// TIA Portal project "Network_1.0" (V15.1) (continued)
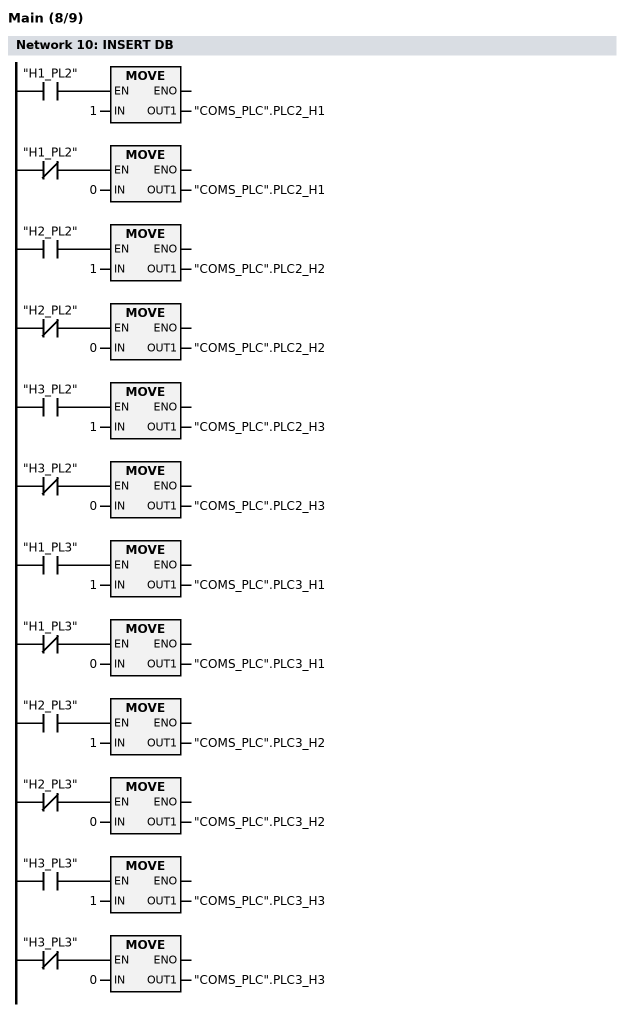
   RUNG wire#powerrail
      Contact( "H1_PL2" )
      Move(in := 1, out1 => "COMS_PLC".PLC2_H1)
   END_RUNG
   RUNG wire#powerrail
      I_Contact( "H1_PL2" )
      Move(in := 0, out1 => "COMS_PLC".PLC2_H1)
   END_RUNG
   RUNG wire#powerrail
      Contact( "H2_PL2" )
      Move(in := 1, out1 => "COMS_PLC".PLC2_H2)
   END_RUNG
   RUNG wire#powerrail
      I_Contact( "H2_PL2" )
      Move(in := 0, out1 => "COMS_PLC".PLC2_H2)
   END_RUNG
   RUNG wire#powerrail
      Contact( "H3_PL2" )
      Move(in := 1, out1 => "COMS_PLC".PLC2_H3)
   END_RUNG
   RUNG wire#powerrail
      I_Contact( "H3_PL2" )
      Move(in := 0, out1 => "COMS_PLC".PLC2_H3)
   END_RUNG
   RUNG wire#powerrail
      Contact( "H1_PL3" )
      Move(in := 1, out1 => "COMS_PLC".PLC3_H1)
   END_RUNG
   RUNG wire#powerrail
      I_Contact( "H1_PL3" )
      Move(in := 0, out1 => "COMS_PLC".PLC3_H1)
   END_RUNG
   RUNG wire#powerrail
      Contact( "H2_PL3" )
      Move(in := 1, out1 => "COMS_PLC".PLC3_H2)
   END_RUNG
   RUNG wire#powerrail
      I_Contact( "H2_PL3" )
      Move(in := 0, out1 => "COMS_PLC".PLC3_H2)
   END_RUNG
   RUNG wire#powerrail
      Contact( "H3_PL3" )
      Move(in := 1, out1 => "COMS_PLC".PLC3_H3)
   END_RUNG
   RUNG wire#powerrail
      I_Contact( "H3_PL3" )
      Move(in := 0, out1 => "COMS_PLC".PLC3_H3)
   END_RUNG
   // the same network as SCL:
   IF "H1_PL2" THEN "COMS_PLC".PLC2_H1 := 1; END_IF;
   IF NOT "H1_PL2" THEN "COMS_PLC".PLC2_H1 := 0; END_IF;
   IF "H2_PL2" THEN "COMS_PLC".PLC2_H2 := 1; END_IF;
   IF NOT "H2_PL2" THEN "COMS_PLC".PLC2_H2 := 0; END_IF;
   IF "H3_PL2" THEN "COMS_PLC".PLC2_H3 := 1; END_IF;
   IF NOT "H3_PL2" THEN "COMS_PLC".PLC2_H3 := 0; END_IF;
   IF "H1_PL3" THEN "COMS_PLC".PLC3_H1 := 1; END_IF;
   IF NOT "H1_PL3" THEN "COMS_PLC".PLC3_H1 := 0; END_IF;
   IF "H2_PL3" THEN "COMS_PLC".PLC3_H2 := 1; END_IF;
   IF NOT "H2_PL3" THEN "COMS_PLC".PLC3_H2 := 0; END_IF;
   IF "H3_PL3" THEN "COMS_PLC".PLC3_H3 := 1; END_IF;
   IF NOT "H3_PL3" THEN "COMS_PLC".PLC3_H3 := 0; END_IF;
END_REGION

REGION Network 11: GET
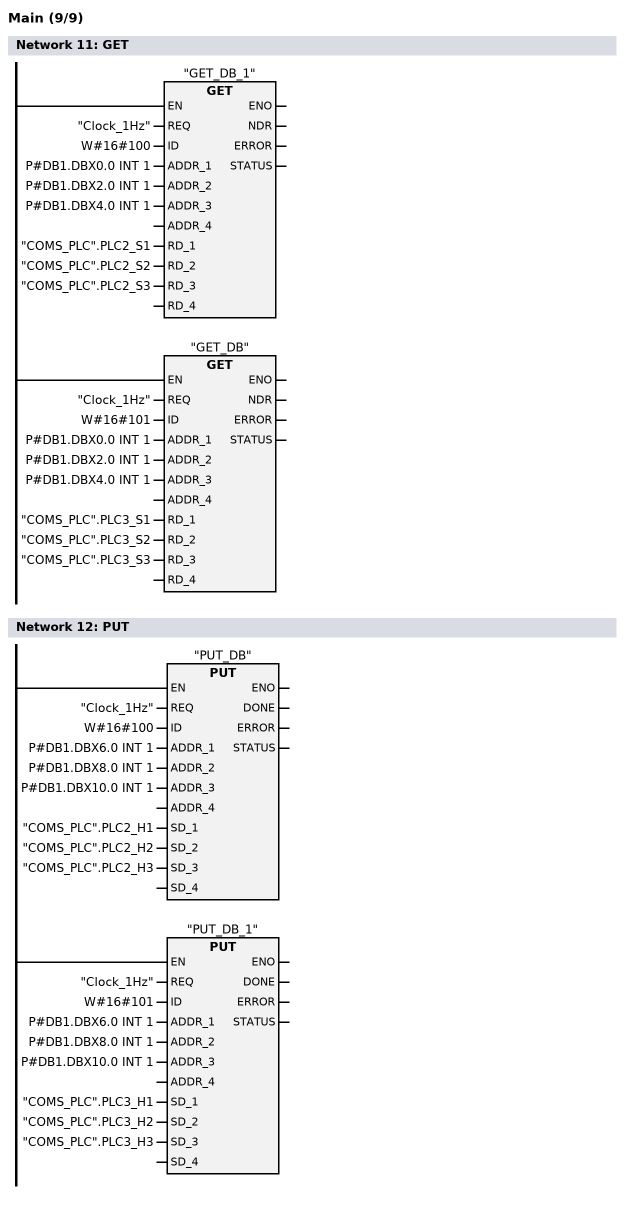
   "GET_DB_1"(REQ := "Clock_1Hz",   // GET
              ID := W#16#100,
              ADDR_1 := P#DB1.DBX0.0 INT 1,
              ADDR_2 := P#DB1.DBX2.0 INT 1,
              ADDR_3 := P#DB1.DBX4.0 INT 1,
              RD_1 := "COMS_PLC".PLC2_S1,
              RD_2 := "COMS_PLC".PLC2_S2,
              RD_3 := "COMS_PLC".PLC2_S3);
   "GET_DB"(REQ := "Clock_1Hz",   // GET
            ID := W#16#101,
            ADDR_1 := P#DB1.DBX0.0 INT 1,
            ADDR_2 := P#DB1.DBX2.0 INT 1,
            ADDR_3 := P#DB1.DBX4.0 INT 1,
            RD_1 := "COMS_PLC".PLC3_S1,
            RD_2 := "COMS_PLC".PLC3_S2,
            RD_3 := "COMS_PLC".PLC3_S3);
END_REGION

REGION Network 12: PUT
   "PUT_DB"(REQ := "Clock_1Hz",   // PUT
            ID := W#16#100,
            ADDR_1 := P#DB1.DBX6.0 INT 1,
            ADDR_2 := P#DB1.DBX8.0 INT 1,
            ADDR_3 := P#DB1.DBX10.0 INT 1,
            SD_1 := "COMS_PLC".PLC2_H1,
            SD_2 := "COMS_PLC".PLC2_H2,
            SD_3 := "COMS_PLC".PLC2_H3);
   "PUT_DB_1"(REQ := "Clock_1Hz",   // PUT
              ID := W#16#101,
              ADDR_1 := P#DB1.DBX6.0 INT 1,
              ADDR_2 := P#DB1.DBX8.0 INT 1,
              ADDR_3 := P#DB1.DBX10.0 INT 1,
              SD_1 := "COMS_PLC".PLC3_H1,
              SD_2 := "COMS_PLC".PLC3_H2,
              SD_3 := "COMS_PLC".PLC3_H3);
END_REGION
END_ORGANIZATION_BLOCK

// ===== PLC "PLC_2"  CPU 1215C DC/DC/DC =====

VAR_GLOBAL   // PLC tag table "Default tag table"
   "S4_JR" AT %I0.0 : Bool;
   "S3_JR" AT %I0.1 : Bool;
   "H2_JR" AT %Q0.1 : Bool;
   "S2_JR" AT %I0.2 : Bool;
   "S1_JR" AT %I0.3 : Bool;
   "PE_JR" AT %I0.4 : Bool;
   "H1_JR" AT %Q0.2 : Bool;
   "H3_JR" AT %Q0.0 : Bool;
   "Clock_Byte" AT %MB0 : Byte;
   "Clock_10Hz" AT %M0.0 : Bool;
   "Clock_5Hz" AT %M0.1 : Bool;
   "Clock_2.5Hz" AT %M0.2 : Bool;
   "Clock_2Hz" AT %M0.3 : Bool;
   "Clock_1.25Hz" AT %M0.4 : Bool;
   "Clock_1Hz" AT %M0.5 : Bool;
   "Clock_0.625Hz" AT %M0.6 : Bool;
   "Clock_0.5Hz" AT %M0.7 : Bool;
END_VAR

VAR_GLOBAL CONSTANT   // PLC tag table "Default tag table"
   "PLC_2" : Byte := 11;   // 2
END_VAR

DATA_BLOCK "Prueba"   // DB1
{ S7_Optimized_Access := 'FALSE' }
VERSION : 0.1
   VAR
      S1 : Int;
      S2 : Int;
      S3 : Int;
      H1 : Int;
      H2 : Int;
      H3 : Int;
   END_VAR
BEGIN
END_DATA_BLOCK

ORGANIZATION_BLOCK "Main"   // OB1, LAD, ProgramCycle
TITLE = "Main Program Sweep (Cycle)"
{ S7_Optimized_Access := 'TRUE' }
VERSION : 0.1
   VAR_INPUT
      Initial_Call : Bool;   // Initial call of this OB
      Remanence : Bool;   // =True, if remanent data are available
   END_VAR
BEGIN

REGION Network 1: SET DB
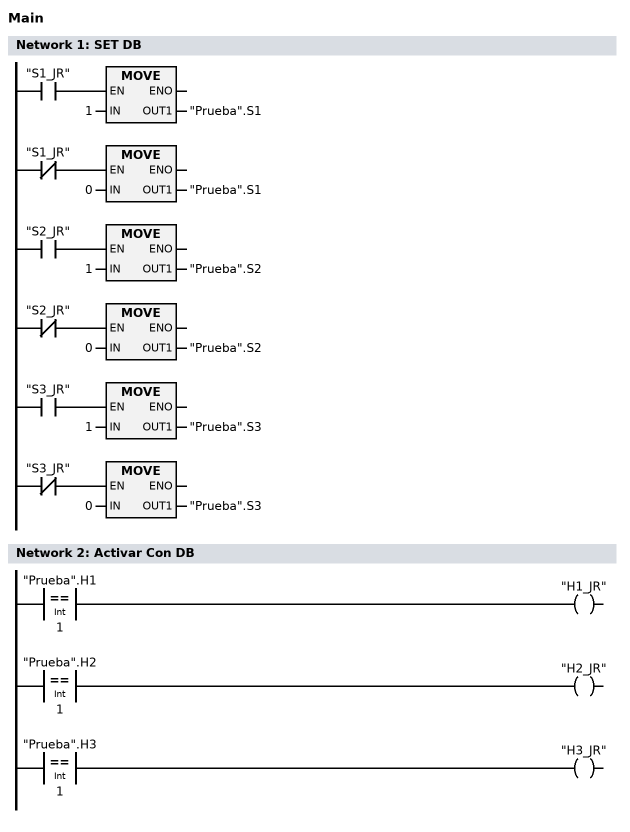
   RUNG wire#powerrail
      Contact( "S1_JR" )
      Move(in := 1, out1 => "Prueba".S1)
   END_RUNG
   RUNG wire#powerrail
      I_Contact( "S1_JR" )
      Move(in := 0, out1 => "Prueba".S1)
   END_RUNG
   RUNG wire#powerrail
      Contact( "S2_JR" )
      Move(in := 1, out1 => "Prueba".S2)
   END_RUNG
   RUNG wire#powerrail
      I_Contact( "S2_JR" )
      Move(in := 0, out1 => "Prueba".S2)
   END_RUNG
   RUNG wire#powerrail
      Contact( "S3_JR" )
      Move(in := 1, out1 => "Prueba".S3)
   END_RUNG
   RUNG wire#powerrail
      I_Contact( "S3_JR" )
      Move(in := 0, out1 => "Prueba".S3)
   END_RUNG
   // the same network as SCL:
   IF "S1_JR" THEN "Prueba".S1 := 1; END_IF;
   IF NOT "S1_JR" THEN "Prueba".S1 := 0; END_IF;
   IF "S2_JR" THEN "Prueba".S2 := 1; END_IF;
   IF NOT "S2_JR" THEN "Prueba".S2 := 0; END_IF;
   IF "S3_JR" THEN "Prueba".S3 := 1; END_IF;
   IF NOT "S3_JR" THEN "Prueba".S3 := 0; END_IF;
END_REGION

REGION Network 2: Activar Con DB
   RUNG wire#powerrail
      { S7_Templates := "SrcType := Int" } EQ_Contact(in1 := "Prueba".H1, in2 := 1)
      Coil( "H1_JR" )
   END_RUNG
   RUNG wire#powerrail
      { S7_Templates := "SrcType := Int" } EQ_Contact(in1 := "Prueba".H2, in2 := 1)
      Coil( "H2_JR" )
   END_RUNG
   RUNG wire#powerrail
      { S7_Templates := "SrcType := Int" } EQ_Contact(in1 := "Prueba".H3, in2 := 1)
      Coil( "H3_JR" )
   END_RUNG
   // the same network as SCL:
   "H1_JR" := "Prueba".H1 = 1;
   "H2_JR" := "Prueba".H2 = 1;
   "H3_JR" := "Prueba".H3 = 1;
END_REGION
END_ORGANIZATION_BLOCK

// ===== PLC "PLC_3"  CPU 1215C DC/DC/DC =====

VAR_GLOBAL   // PLC tag table "Default tag table"
   "H1_FE" AT %Q0.0 : Bool;
   "PE_FE" AT %I0.0 : Bool;
   "S1_FE" AT %I0.1 : Bool;
   "S2_FE" AT %I0.2 : Bool;
   "S3_FE" AT %I0.3 : Bool;
   "H2_FE" AT %Q0.1 : Bool;
   "H3_FE" AT %Q0.2 : Bool;
END_VAR

DATA_BLOCK "Control_PLC3"   // DB1
{ S7_Optimized_Access := 'FALSE' }
VERSION : 0.1
   VAR
      S1 : Int;
      S2 : Int;
      S3 : Int;
      H1 : Int;
      H2 : Int;
      H3 : Int;
   END_VAR
BEGIN
END_DATA_BLOCK

ORGANIZATION_BLOCK "Main"   // OB1, LAD, ProgramCycle
TITLE = "Main Program Sweep (Cycle)"
{ S7_Optimized_Access := 'TRUE' }
VERSION : 0.1
   VAR_INPUT
      Initial_Call : Bool;   // Initial call of this OB
      Remanence : Bool;   // =True, if remanent data are available
   END_VAR
BEGIN

REGION Network 1: SET DB
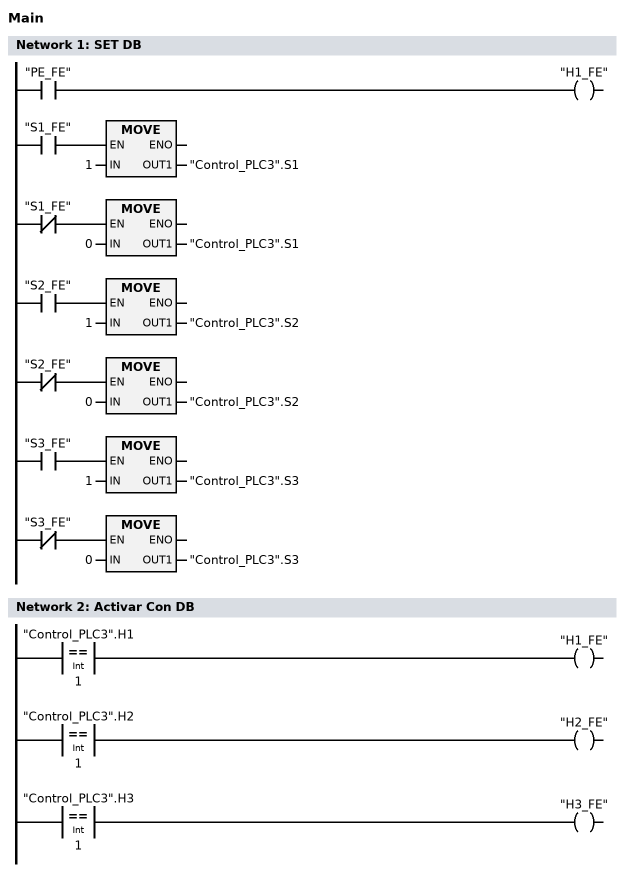
   RUNG wire#powerrail
      Contact( "PE_FE" )
      Coil( "H1_FE" )
   END_RUNG
   RUNG wire#powerrail
      Contact( "S1_FE" )
      Move(in := 1, out1 => "Control_PLC3".S1)
   END_RUNG
   RUNG wire#powerrail
      I_Contact( "S1_FE" )
      Move(in := 0, out1 => "Control_PLC3".S1)
   END_RUNG
   RUNG wire#powerrail
      Contact( "S2_FE" )
      Move(in := 1, out1 => "Control_PLC3".S2)
   END_RUNG
   RUNG wire#powerrail
      I_Contact( "S2_FE" )
      Move(in := 0, out1 => "Control_PLC3".S2)
   END_RUNG
   RUNG wire#powerrail
      Contact( "S3_FE" )
      Move(in := 1, out1 => "Control_PLC3".S3)
   END_RUNG
   RUNG wire#powerrail
      I_Contact( "S3_FE" )
      Move(in := 0, out1 => "Control_PLC3".S3)
   END_RUNG
   // the same network as SCL:
   "H1_FE" := "PE_FE";
   IF "S1_FE" THEN "Control_PLC3".S1 := 1; END_IF;
   IF NOT "S1_FE" THEN "Control_PLC3".S1 := 0; END_IF;
   IF "S2_FE" THEN "Control_PLC3".S2 := 1; END_IF;
   IF NOT "S2_FE" THEN "Control_PLC3".S2 := 0; END_IF;
   IF "S3_FE" THEN "Control_PLC3".S3 := 1; END_IF;
   IF NOT "S3_FE" THEN "Control_PLC3".S3 := 0; END_IF;
END_REGION

REGION Network 2: Activar Con DB
   RUNG wire#powerrail
      { S7_Templates := "SrcType := Int" } EQ_Contact(in1 := "Control_PLC3".H1, in2 := 1)
      Coil( "H1_FE" )
   END_RUNG
   RUNG wire#powerrail
      { S7_Templates := "SrcType := Int" } EQ_Contact(in1 := "Control_PLC3".H2, in2 := 1)
      Coil( "H2_FE" )
   END_RUNG
   RUNG wire#powerrail
      { S7_Templates := "SrcType := Int" } EQ_Contact(in1 := "Control_PLC3".H3, in2 := 1)
      Coil( "H3_FE" )
   END_RUNG
   // the same network as SCL:
   "H1_FE" := "Control_PLC3".H1 = 1;
   "H2_FE" := "Control_PLC3".H2 = 1;
   "H3_FE" := "Control_PLC3".H3 = 1;
END_REGION
END_ORGANIZATION_BLOCK

(* ===== HMI "HMI_RT_1" =====
system functions are stored by id; their names below are inferred from use
connection "HMI_Connection_1": ETHERNET, SMART_S7_1500_OMS

HMI tags "Default tag table"
   "Tag_ScreenNumber" : UInt, internal
   "S1" : Bool = PLC S1_HM1 AT %M3.0, 100 ms
   "S2" : Bool = PLC S2_HM1 AT %M3.1, 100 ms
   "S3" : Bool = PLC S3_HM1 AT %M3.2, 100 ms
   "H1_HM1" : Bool = PLC H1_HM1 AT %M6.3, 100 ms
   "H2_HM1" : Bool = PLC H2_HM1 AT %M6.4, 100 ms
   "H3_HM1" : Bool = PLC H3_HM1 AT %M6.5, 100 ms
   "Selector" : UInt = PLC Selector_HMI_1 AT %MW8, 100 ms

text list "PLC_SELECTOR": 1 'Betsy'; 2 'JR'; 3 'Fer'

Template "Template_1" 480x272
   Button "Exit" at 388,227 size 63x44; TextOff 'Exit'; PictureOff "ExitRuntime_KTP400_Basic_PN_TR"; PictureOn "ExitRuntime_KTP400_Basic_PN_TR"
      on Release: StopRuntime(0)
   Button "Log on" at 268,227 size 63x44; TextOff 'Log on'; PictureOff "Login_KTP400_Basic_PN_TR"; PictureOn "Login_KTP400_Basic_PN_TR"
      on Release: function_a2a04561()
   Button "Alarms" at 148,227 size 63x44; TextOff 'Alarms'; PictureOff "AlarmDisplay_KTP400_Basic_PN_TR"; PictureOn "AlarmDisplay_KTP400_Basic_PN_TR"
      on Release: function_ef3f5d25("Alarm window_Unacknowledged", -1)
   Button "Start screen" at 28,227 size 63x44; TextOff 'Start screen'; PictureOff "NavigateHome_KTP400_Basic_PN_TR"; PictureOn "NavigateHome_KTP400_Basic_PN_TR"
      on Release: ActivateScreen("Root screen", 0)
   SymbolicIOField "Symbolic_IO_Field_Screen" at 162,8 size 231x29; TextOff '0'; TextOn '1'; TextList "TextList_ScreenNames"
      ProcessValue <- "Tag_ScreenNumber"
      on Change: ActivateScreenByNumber("Tag_ScreenNumber", 0)
   DateTimeField "HmiScreenItemData" at 395,22 size 85x22
   DateTimeField "HmiScreenItemData_1" at 395,0 size 85x22
   GraphicView "Logo" at 0,0 size 160x45; Picture "Logo of HMI_1"

screen "Root screen" 480x272, template "Template_1"
   on GenerateScreen: SetTag("Tag_ScreenNumber", 1)
   Button "Button_1" at 169,112 size 146x61; TextOff 'LED CONTROL'
      on Click: ActivateScreen("Led_control", 8)

screen "SIMATIC PLC system diagnostics" 480x272, template "Template_1"
   on GenerateScreen: SetTag("Tag_ScreenNumber", 3)
   SysDiagControl "HmiScreenItemData" at 1,77 size 476x143
   Button "Back" at 1,46 size 157x30; TextOff 'Back'
      on Release: ActivateScreen("Root screen", 0)

screen "Project information" 480x272, template "Template_1"
   on GenerateScreen: SetTag("Tag_ScreenNumber", 4)
   TextField "HmiScreenItemData" at 4,78 size 184x20; Text 'Project name:'
   TextField "HmiScreenItemData_1" at 192,78 size 284x20; Text 'Network_1'
   TextField "HmiScreenItemData_2" at 4,99 size 184x20; Text 'Created on:'
   TextField "HmiScreenItemData_3" at 192,99 size 284x20; Text '3/10/2025 2:35:17 PM'
   TextField "HmiScreenItemData_4" at 4,120 size 184x20; Text 'Author:'
   TextField "HmiScreenItemData_5" at 192,120 size 284x20; Text '192072'
   TextField "HmiScreenItemData_6" at 4,141 size 184x20; Text 'Description:'
   TextField "HmiScreenItemData_7" at 192,141 size 284x20; Text '(not configured)'
   Button "Back" at 1,46 size 157x30; TextOff 'Back'
      on Release: ActivateScreen("Root screen", 0)

screen "System information" 480x272, template "Template_1"
   on GenerateScreen: SetTag("Tag_ScreenNumber", 6)
   TextField "HmiScreenItemData" at 4,78 size 184x20; Text 'HMI device type:'
   TextField "HmiScreenItemData_1" at 192,78 size 284x20; Text 'KTP400 Basic+ PN 15.1.0.0'
   TextField "HmiScreenItemData_2" at 4,99 size 184x20; Text 'Connection:'
   TextField "HmiScreenItemData_3" at 192,99 size 284x20; Text '(not configured)'
   TextField "HmiScreenItemData_4" at 4,120 size 184x20; Text 'PLC:'
   TextField "HmiScreenItemData_5" at 192,120 size 284x20; Text '<PLC>'
   Button "Back" at 1,46 size 157x30; TextOff 'Back'
      on Release: ActivateScreen("Root screen", 0)

screen "Led_control" 480x272
   Circle "Circle_1" at 58,80 size 86x86
      Appearance <- "H1_HM1"
   Circle "Circle_2" at 203,80 size 86x86
      Appearance <- "H2_HM1"
   Circle "Circle_3" at 348,80 size 86x86
      Appearance <- "H3_HM1"
   GraphicView "Graphic view_1" at 0,6 size 148x37; Picture "Logo of HMI_3"
   SymbolicIOField "Symbolic I/O field_1" at 321,5 size 152x35; TextOff '0'; TextOn '1'; TextList "PLC_SELECTOR"
      ProcessValue <- "Selector"
   Button "Button_1" at 47,215 size 102x28; TextOff 'S1'
      on Release: SetTag("S1", 0)
      on Press: SetTag("S1", 1)
   Button "Button_2" at 195,215 size 102x28; TextOff 'S2'
      on Press: SetTag("S2", 1)
      on Release: SetTag("S2", 0)
   Button "Button_3" at 341,215 size 102x28; TextOff 'S3'
      on Press: SetTag("S3", 1)
      on Release: SetTag("S3", 0)
   Button "Button_4" at 203,6 size 96x32; TextOff 'Back'
      on Click: function_efd93a16()
*)

(* ===== HMI "HMI_RT_2" =====
system functions are stored by id; their names below are inferred from use
connection "HMI_Connection_2": ETHERNET, SMART_S7_1500_OMS

HMI tags "Default tag table"
   "Tag_ScreenNumber" : UInt, internal
   "H1_HM2" : Bool = PLC H1_HM2 AT %M6.6, 100 ms
   "H2_HM2" : Bool = PLC H2_HM2 AT %M6.7, 100 ms
   "H3_HM2" : Bool = PLC H3_HM2 AT %M7.0, 100 ms
   "S1" : Bool = PLC S1_HM2 AT %M3.3, 100 ms
   "S2" : Bool = PLC S2_HM2 AT %M3.4, 100 ms
   "S3" : Bool = PLC S3_HM2 AT %M3.5, 100 ms
   "Selector" : UInt = PLC Selector_HMI_2 AT %MW10, 100 ms

text list "PLC_SELECTOR": 1 'Betsy'; 2 'JR'; 3 'Fer'

Template "Template_1" 480x272
   Button "Exit" at 388,227 size 63x44; TextOff 'Exit'; PictureOff "ExitRuntime_KTP400_Basic_PN_TR"; PictureOn "ExitRuntime_KTP400_Basic_PN_TR"
      on Release: StopRuntime(0)
   Button "Log on" at 268,227 size 63x44; TextOff 'Log on'; PictureOff "Login_KTP400_Basic_PN_TR"; PictureOn "Login_KTP400_Basic_PN_TR"
      on Release: function_a2a04561()
   Button "Alarms" at 148,227 size 63x44; TextOff 'Alarms'; PictureOff "AlarmDisplay_KTP400_Basic_PN_TR"; PictureOn "AlarmDisplay_KTP400_Basic_PN_TR"
      on Release: function_ef3f5d25("Alarm window_Unacknowledged", -1)
   Button "Start screen" at 28,227 size 63x44; TextOff 'Start screen'; PictureOff "NavigateHome_KTP400_Basic_PN_TR"; PictureOn "NavigateHome_KTP400_Basic_PN_TR"
      on Release: ActivateScreen("Root screen", 0)
   SymbolicIOField "Symbolic_IO_Field_Screen" at 162,8 size 231x29; TextOff '0'; TextOn '1'; TextList "TextList_ScreenNames"
      ProcessValue <- "Tag_ScreenNumber"
      on Change: ActivateScreenByNumber("Tag_ScreenNumber", 0)
   DateTimeField "HmiScreenItemData" at 395,22 size 85x22
   DateTimeField "HmiScreenItemData_1" at 395,0 size 85x22
   GraphicView "Logo" at 0,0 size 160x45; Picture "Logo of HMI_2"

screen "System screens" 480x272, template "Template_1"
   on GenerateScreen: SetTag("Tag_ScreenNumber", 2)
   TextField "HmiScreenItemData" at 48,122 size 384x22; Text 'System screens'
   Button "Back" at 1,46 size 157x30; TextOff 'Back'
      on Release: ActivateScreen("Root screen", 0)
   Button "SIMATIC PLC system diagnostics" at 1,77 size 157x30; TextOff 'SIMATIC PLC syst...'
      on Release: ActivateScreen("SIMATIC PLC system diagnostics", 0)
   Button "Project information" at 1,108 size 157x30; TextOff 'Project information'
      on Release: ActivateScreen("Project information", 0)
   Button "User administration" at 1,139 size 157x30; TextOff 'User administration'
      on Release: ActivateScreen("User administration", 0)
   Button "System information" at 1,170 size 157x30; TextOff 'System information'
      on Release: ActivateScreen("System information", 0)
   Button "Different jobs" at 159,46 size 157x30; TextOff 'Different jobs'
      on Release: ActivateScreen("Different jobs", 0)

screen "SIMATIC PLC system diagnostics" 480x272, template "Template_1"
   on GenerateScreen: SetTag("Tag_ScreenNumber", 3)
   SysDiagControl "HmiScreenItemData" at 1,77 size 476x143
   Button "Back" at 1,46 size 157x30; TextOff 'Back'
      on Release: ActivateScreen("System screens", 0)

screen "Project information" 480x272, template "Template_1"
   on GenerateScreen: SetTag("Tag_ScreenNumber", 4)
   TextField "HmiScreenItemData" at 4,78 size 184x20; Text 'Project name:'
   TextField "HmiScreenItemData_1" at 192,78 size 284x20; Text 'Network_1'
   TextField "HmiScreenItemData_2" at 4,99 size 184x20; Text 'Created on:'
   TextField "HmiScreenItemData_3" at 192,99 size 284x20; Text '3/10/2025 2:35:17 PM'
   TextField "HmiScreenItemData_4" at 4,120 size 184x20; Text 'Author:'
   TextField "HmiScreenItemData_5" at 192,120 size 284x20; Text '192072'
   TextField "HmiScreenItemData_6" at 4,141 size 184x20; Text 'Description:'
   TextField "HmiScreenItemData_7" at 192,141 size 284x20; Text '(not configured)'
   Button "Back" at 1,46 size 157x30; TextOff 'Back'
      on Release: ActivateScreen("System screens", 0)

screen "User administration" 480x272, template "Template_1"
   on GenerateScreen: SetTag("Tag_ScreenNumber", 5)
   UserView "HmiScreenItemData" at 1,77 size 476x143
   Button "Back" at 1,46 size 157x30; TextOff 'Back'
      on Release: ActivateScreen("System screens", 0)

screen "System information" 480x272, template "Template_1"
   on GenerateScreen: SetTag("Tag_ScreenNumber", 6)
   TextField "HmiScreenItemData" at 4,78 size 184x20; Text 'HMI device type:'
   TextField "HmiScreenItemData_1" at 192,78 size 284x20; Text 'KTP400 Basic+ PN 15.1.0.0'
   TextField "HmiScreenItemData_2" at 4,99 size 184x20; Text 'Connection:'
   TextField "HmiScreenItemData_3" at 192,99 size 284x20; Text '(not configured)'
   TextField "HmiScreenItemData_4" at 4,120 size 184x20; Text 'PLC:'
   TextField "HmiScreenItemData_5" at 192,120 size 284x20; Text '<PLC>'
   Button "Back" at 1,46 size 157x30; TextOff 'Back'
      on Release: ActivateScreen("System screens", 0)

screen "Different jobs" 480x272, template "Template_1"
   on GenerateScreen: SetTag("Tag_ScreenNumber", 7)
   Button "Online" at 1,77 size 157x30; TextOff 'Online'
      on Release: function_bb44b551(0)
   Button "Offline" at 1,108 size 157x30; TextOff 'Offline'
      on Release: function_bb44b551(1)
   Button "Transfer" at 1,139 size 157x30; TextOff 'Transfer'
      on Release: function_bb44b551(2)
   Button "Toggle language" at 1,170 size 157x30; TextOff 'Toggle language'
      on Release: function_fb9197e8(-1)
   Button "Stop Runtime" at 159,77 size 157x30; TextOff 'Stop Runtime'
      on Release: StopRuntime(0)
   Button "Back" at 1,46 size 157x30; TextOff 'Back'
      on Release: ActivateScreen("System screens", 0)

screen "Root screen" 480x272, template "Template_1"
   on GenerateScreen: SetTag("Tag_ScreenNumber", 1)
   Button "Button_1" at 169,112 size 146x61; TextOff 'LED CONTROL'
      on Click: ActivateScreen("Led_control", 8)

screen "Led_control" 480x272
   Circle "Circle_1" at 58,80 size 86x86
      Appearance <- "H1_HM2"
   Circle "Circle_2" at 203,80 size 86x86
      Appearance <- "H2_HM2"
   Circle "Circle_3" at 348,80 size 86x86
      Appearance <- "H3_HM2"
   GraphicView "Graphic view_1" at 0,6 size 148x37; Picture "Logo of HMI_3"
   SymbolicIOField "Symbolic I/O field_1" at 321,5 size 152x35; TextOn '1'; TextOff '0'; TextList "PLC_SELECTOR"
      ProcessValue <- "Selector"
   Button "Button_1" at 47,215 size 102x28; TextOff 'S1'
      on Release: SetTag("S1", 0)
      on Press: SetTag("S1", 1)
   Button "Button_2" at 195,215 size 102x28; TextOff 'S2'
      on Release: SetTag("S2", 0)
      on Press: SetTag("S2", 1)
   Button "Button_3" at 341,215 size 102x28; TextOff 'S3'
      on Release: SetTag("S3", 0)
      on Press: SetTag("S3", 1)
   Button "Button_4" at 203,6 size 96x32; TextOff 'Back'
      on Click: function_efd93a16()
*)

(* ===== HMI "HMI_RT_3" =====
system functions are stored by id; their names below are inferred from use
connection "HMI_Connection_4": ETHERNET, SMART_S7_1500_OMS

HMI tags "Default tag table"
   "H1_HM2" : Bool = PLC H1_HM3 AT %M7.1, 100 ms
   "H2_HM2" : Bool = PLC H2_HM3 AT %M7.2, 100 ms
   "H3_HM2" : Bool = PLC H3_HM3 AT %M7.3, 100 ms
   "S1" : Bool = PLC S1_HM3 AT %M3.6, 100 ms
   "S2" : Bool = PLC S2_HM3 AT %M3.7, 100 ms
   "S3" : Bool = PLC S3_HM3 AT %M4.0, 100 ms
   "Tag_ScreenNumber" : UInt, internal
   "Selector" : UInt = PLC Selector_HMI_3 AT %MW12, 100 ms

text list "PLC_SELECTOR": 1 'Betsy'; 2 'JR'; 3 'Fer'

Template "Template_1" 480x272
   Button "Exit" at 388,227 size 63x44; TextOff 'Exit'; PictureOff "ExitRuntime_KTP400_Basic_PN_TR"; PictureOn "ExitRuntime_KTP400_Basic_PN_TR"
      on Release: StopRuntime(0)
   Button "Log on" at 268,227 size 63x44; TextOff 'Log on'; PictureOff "Login_KTP400_Basic_PN_TR"; PictureOn "Login_KTP400_Basic_PN_TR"
      on Release: function_a2a04561()
   Button "Alarms" at 148,227 size 63x44; TextOff 'Alarms'; PictureOff "AlarmDisplay_KTP400_Basic_PN_TR"; PictureOn "AlarmDisplay_KTP400_Basic_PN_TR"
      on Release: function_ef3f5d25("Alarm window_Unacknowledged", -1)
   Button "Start screen" at 28,227 size 63x44; TextOff 'Start screen'; PictureOff "NavigateHome_KTP400_Basic_PN_TR"; PictureOn "NavigateHome_KTP400_Basic_PN_TR"
      on Release: ActivateScreen("Root screen", 0)
   SymbolicIOField "Symbolic_IO_Field_Screen" at 162,8 size 231x29; TextOff '0'; TextOn '1'; TextList "TextList_ScreenNames"
      on Change: ActivateScreenByNumber("Tag_ScreenNumber", 0)
      ProcessValue <- "Tag_ScreenNumber"
   DateTimeField "HmiScreenItemData" at 395,22 size 85x22
   DateTimeField "HmiScreenItemData_1" at 395,0 size 85x22
   GraphicView "Logo" at 0,0 size 160x45; Picture "Logo of HMI_3"

screen "System screens" 480x272, template "Template_1"
   on GenerateScreen: SetTag("Tag_ScreenNumber", 2)
   TextField "HmiScreenItemData" at 48,122 size 384x22; Text 'System screens'
   Button "Back" at 1,46 size 157x30; TextOff 'Back'
      on Release: ActivateScreen("Root screen", 0)
   Button "SIMATIC PLC system diagnostics" at 1,77 size 157x30; TextOff 'SIMATIC PLC syst...'
      on Release: ActivateScreen("SIMATIC PLC system diagnostics", 0)
   Button "Project information" at 1,108 size 157x30; TextOff 'Project information'
      on Release: ActivateScreen("Project information", 0)
   Button "User administration" at 1,139 size 157x30; TextOff 'User administration'
      on Release: ActivateScreen("User administration", 0)
   Button "System information" at 1,170 size 157x30; TextOff 'System information'
      on Release: ActivateScreen("System information", 0)
   Button "Different jobs" at 159,46 size 157x30; TextOff 'Different jobs'
      on Release: ActivateScreen("Different jobs", 0)

screen "SIMATIC PLC system diagnostics" 480x272, template "Template_1"
   on GenerateScreen: SetTag("Tag_ScreenNumber", 3)
   SysDiagControl "HmiScreenItemData" at 1,77 size 476x143
   Button "Back" at 1,46 size 157x30; TextOff 'Back'
      on Release: ActivateScreen("System screens", 0)

screen "Project information" 480x272, template "Template_1"
   on GenerateScreen: SetTag("Tag_ScreenNumber", 4)
   TextField "HmiScreenItemData" at 4,78 size 184x20; Text 'Project name:'
   TextField "HmiScreenItemData_1" at 192,78 size 284x20; Text 'Network_1'
   TextField "HmiScreenItemData_2" at 4,99 size 184x20; Text 'Created on:'
   TextField "HmiScreenItemData_3" at 192,99 size 284x20; Text '3/10/2025 2:35:17 PM'
   TextField "HmiScreenItemData_4" at 4,120 size 184x20; Text 'Author:'
   TextField "HmiScreenItemData_5" at 192,120 size 284x20; Text '192072'
   TextField "HmiScreenItemData_6" at 4,141 size 184x20; Text 'Description:'
   TextField "HmiScreenItemData_7" at 192,141 size 284x20; Text '(not configured)'
   Button "Back" at 1,46 size 157x30; TextOff 'Back'
      on Release: ActivateScreen("System screens", 0)

screen "User administration" 480x272, template "Template_1"
   on GenerateScreen: SetTag("Tag_ScreenNumber", 5)
   UserView "HmiScreenItemData" at 1,77 size 476x143
   Button "Back" at 1,46 size 157x30; TextOff 'Back'
      on Release: ActivateScreen("System screens", 0)

screen "System information" 480x272, template "Template_1"
   on GenerateScreen: SetTag("Tag_ScreenNumber", 6)
   TextField "HmiScreenItemData" at 4,78 size 184x20; Text 'HMI device type:'
   TextField "HmiScreenItemData_1" at 192,78 size 284x20; Text 'KTP400 Basic+ PN 15.1.0.0'
   TextField "HmiScreenItemData_2" at 4,99 size 184x20; Text 'Connection:'
   TextField "HmiScreenItemData_3" at 192,99 size 284x20; Text '(not configured)'
   TextField "HmiScreenItemData_4" at 4,120 size 184x20; Text 'PLC:'
   TextField "HmiScreenItemData_5" at 192,120 size 284x20; Text '<PLC>'
   Button "Back" at 1,46 size 157x30; TextOff 'Back'
      on Release: ActivateScreen("System screens", 0)

screen "Different jobs" 480x272, template "Template_1"
   on GenerateScreen: SetTag("Tag_ScreenNumber", 7)
   Button "Online" at 1,77 size 157x30; TextOff 'Online'
      on Release: function_bb44b551(0)
   Button "Offline" at 1,108 size 157x30; TextOff 'Offline'
      on Release: function_bb44b551(1)
   Button "Transfer" at 1,139 size 157x30; TextOff 'Transfer'
      on Release: function_bb44b551(2)
   Button "Toggle language" at 1,170 size 157x30; TextOff 'Toggle language'
      on Release: function_fb9197e8(-1)
   Button "Stop Runtime" at 159,77 size 157x30; TextOff 'Stop Runtime'
      on Release: StopRuntime(0)
   Button "Back" at 1,46 size 157x30; TextOff 'Back'
      on Release: ActivateScreen("System screens", 0)

screen "Root screen" 480x272, template "Template_1"
   on GenerateScreen: SetTag("Tag_ScreenNumber", 1)
   Button "Button_1" at 169,112 size 146x61; TextOff 'LED CONTROL'
      on Click: ActivateScreen("Led_control", 8)

screen "Led_control" 480x272
   Circle "Circle_1" at 58,80 size 86x86
      Appearance <- "H1_HM2"
   Circle "Circle_2" at 203,80 size 86x86
      Appearance <- "H2_HM2"
   Circle "Circle_3" at 348,80 size 86x86
      Appearance <- "H3_HM2"
   GraphicView "Graphic view_1" at 0,6 size 148x37; Picture "Logo of HMI_3"
   SymbolicIOField "Symbolic I/O field_1" at 321,5 size 152x35; TextOn '1'; TextOff '0'; TextList "PLC_SELECTOR"
      ProcessValue <- "Selector"
   Button "Button_1" at 47,215 size 102x28; TextOff 'S1'
      on Release: SetTag("S1", 0)
      on Press: SetTag("S1", 1)
   Button "Button_2" at 195,215 size 102x28; TextOff 'S2'
      on Release: SetTag("S2", 0)
      on Press: SetTag("S2", 1)
   Button "Button_3" at 341,215 size 102x28; TextOff 'S3'
      on Release: SetTag("S3", 0)
      on Press: SetTag("S3", 1)
   Button "Button_4" at 203,6 size 96x32; TextOff 'Back'
      on Click: function_efd93a16()
*)